HMI tags "DB_SDC_ERROR_STAT_EMS052"
   "DB_SDC_ERRORS_STAT_ER_AKT[52].ER_TRIGER" : Word = PLC DB_SDC_ERRORS_STAT.ER_AKT[52].ER_TRIGER AT %DB3724.DBW31386, 1 s
   "DB_SDC_ERRORS_STAT_ER_AKT[52].ER_STAT[1].DRIVE_POS" : DInt = PLC DB_SDC_ERRORS_STAT.ER_AKT[52].ER_STAT[1].DRIVE_POS AT %DB3724.DBD31392, 1 s
   "DB_SDC_ERRORS_STAT_ER_AKT[52].ER_STAT[1].ERROR" : Int = PLC DB_SDC_ERRORS_STAT.ER_AKT[52].ER_STAT[1].ERROR AT %DB3724.DBW31398, 1 s
   "DB_SDC_ERRORS_STAT_ER_AKT[52].ER_STAT[2].DRIVE_POS" : DInt = PLC DB_SDC_ERRORS_STAT.ER_AKT[52].ER_STAT[2].DRIVE_POS AT %DB3724.DBD31408, 1 s
   "DB_SDC_ERRORS_STAT_ER_AKT[52].ER_STAT[2].ERROR" : Int = PLC DB_SDC_ERRORS_STAT.ER_AKT[52].ER_STAT[2].ERROR AT %DB3724.DBW31414, 1 s
   "DB_SDC_ERRORS_STAT_ER_AKT[52].ER_STAT[3].DRIVE_POS" : DInt = PLC DB_SDC_ERRORS_STAT.ER_AKT[52].ER_STAT[3].DRIVE_POS AT %DB3724.DBD31424, 1 s
   "DB_SDC_ERRORS_STAT_ER_AKT[52].ER_STAT[3].ERROR" : Int = PLC DB_SDC_ERRORS_STAT.ER_AKT[52].ER_STAT[3].ERROR AT %DB3724.DBW31430, 1 s
   "DB_SDC_ERRORS_STAT_ER_AKT[52].ER_STAT[4].DRIVE_POS" : DInt = PLC DB_SDC_ERRORS_STAT.ER_AKT[52].ER_STAT[4].DRIVE_POS AT %DB3724.DBD31440, 1 s
   "DB_SDC_ERRORS_STAT_ER_AKT[52].ER_STAT[4].ERROR" : Int = PLC DB_SDC_ERRORS_STAT.ER_AKT[52].ER_STAT[4].ERROR AT %DB3724.DBW31446, 1 s

HMI tags "DB_SDC_ERROR_STAT_EMS053"
   "DB_SDC_ERRORS_STAT_ER_AKT[53].ER_TRIGER" : Word = PLC DB_SDC_ERRORS_STAT.ER_AKT[53].ER_TRIGER AT %DB3724.DBW31452, 1 s
   "DB_SDC_ERRORS_STAT_ER_AKT[53].ER_STAT[1].DRIVE_POS" : DInt = PLC DB_SDC_ERRORS_STAT.ER_AKT[53].ER_STAT[1].DRIVE_POS AT %DB3724.DBD31458, 1 s
   "DB_SDC_ERRORS_STAT_ER_AKT[53].ER_STAT[1].ERROR" : Int = PLC DB_SDC_ERRORS_STAT.ER_AKT[53].ER_STAT[1].ERROR AT %DB3724.DBW31464, 1 s
   "DB_SDC_ERRORS_STAT_ER_AKT[53].ER_STAT[2].DRIVE_POS" : DInt = PLC DB_SDC_ERRORS_STAT.ER_AKT[53].ER_STAT[2].DRIVE_POS AT %DB3724.DBD31474, 1 s
   "DB_SDC_ERRORS_STAT_ER_AKT[53].ER_STAT[2].ERROR" : Int = PLC DB_SDC_ERRORS_STAT.ER_AKT[53].ER_STAT[2].ERROR AT %DB3724.DBW31480, 1 s
   "DB_SDC_ERRORS_STAT_ER_AKT[53].ER_STAT[3].DRIVE_POS" : DInt = PLC DB_SDC_ERRORS_STAT.ER_AKT[53].ER_STAT[3].DRIVE_POS AT %DB3724.DBD31490, 1 s
   "DB_SDC_ERRORS_STAT_ER_AKT[53].ER_STAT[3].ERROR" : Int = PLC DB_SDC_ERRORS_STAT.ER_AKT[53].ER_STAT[3].ERROR AT %DB3724.DBW31496, 1 s
   "DB_SDC_ERRORS_STAT_ER_AKT[53].ER_STAT[4].DRIVE_POS" : DInt = PLC DB_SDC_ERRORS_STAT.ER_AKT[53].ER_STAT[4].DRIVE_POS AT %DB3724.DBD31506, 1 s
   "DB_SDC_ERRORS_STAT_ER_AKT[53].ER_STAT[4].ERROR" : Int = PLC DB_SDC_ERRORS_STAT.ER_AKT[53].ER_STAT[4].ERROR AT %DB3724.DBW31512, 1 s

HMI tags "DB_SDC_ERROR_STAT_EMS054"
   "DB_SDC_ERRORS_STAT_ER_AKT[54].ER_TRIGER" : Word = PLC DB_SDC_ERRORS_STAT.ER_AKT[54].ER_TRIGER AT %DB3724.DBW31518, 1 s
   "DB_SDC_ERRORS_STAT_ER_AKT[54].ER_STAT[1].DRIVE_POS" : DInt = PLC DB_SDC_ERRORS_STAT.ER_AKT[54].ER_STAT[1].DRIVE_POS AT %DB3724.DBD31524, 1 s
   "DB_SDC_ERRORS_STAT_ER_AKT[54].ER_STAT[1].ERROR" : Int = PLC DB_SDC_ERRORS_STAT.ER_AKT[54].ER_STAT[1].ERROR AT %DB3724.DBW31530, 1 s
   "DB_SDC_ERRORS_STAT_ER_AKT[54].ER_STAT[2].DRIVE_POS" : DInt = PLC DB_SDC_ERRORS_STAT.ER_AKT[54].ER_STAT[2].DRIVE_POS AT %DB3724.DBD31540, 1 s
   "DB_SDC_ERRORS_STAT_ER_AKT[54].ER_STAT[2].ERROR" : Int = PLC DB_SDC_ERRORS_STAT.ER_AKT[54].ER_STAT[2].ERROR AT %DB3724.DBW31546, 1 s
   "DB_SDC_ERRORS_STAT_ER_AKT[54].ER_STAT[3].DRIVE_POS" : DInt = PLC DB_SDC_ERRORS_STAT.ER_AKT[54].ER_STAT[3].DRIVE_POS AT %DB3724.DBD31556, 1 s
   "DB_SDC_ERRORS_STAT_ER_AKT[54].ER_STAT[3].ERROR" : Int = PLC DB_SDC_ERRORS_STAT.ER_AKT[54].ER_STAT[3].ERROR AT %DB3724.DBW31562, 1 s
   "DB_SDC_ERRORS_STAT_ER_AKT[54].ER_STAT[4].DRIVE_POS" : DInt = PLC DB_SDC_ERRORS_STAT.ER_AKT[54].ER_STAT[4].DRIVE_POS AT %DB3724.DBD31572, 1 s
   "DB_SDC_ERRORS_STAT_ER_AKT[54].ER_STAT[4].ERROR" : Int = PLC DB_SDC_ERRORS_STAT.ER_AKT[54].ER_STAT[4].ERROR AT %DB3724.DBW31578, 1 s

HMI tags "DB_SDC_ERROR_STAT_EMS055"
   "DB_SDC_ERRORS_STAT_ER_AKT[55].ER_TRIGER" : Word = PLC DB_SDC_ERRORS_STAT.ER_AKT[55].ER_TRIGER AT %DB3724.DBW31584, 1 s
   "DB_SDC_ERRORS_STAT_ER_AKT[55].ER_STAT[1].DRIVE_POS" : DInt = PLC DB_SDC_ERRORS_STAT.ER_AKT[55].ER_STAT[1].DRIVE_POS AT %DB3724.DBD31590, 1 s
   "DB_SDC_ERRORS_STAT_ER_AKT[55].ER_STAT[1].ERROR" : Int = PLC DB_SDC_ERRORS_STAT.ER_AKT[55].ER_STAT[1].ERROR AT %DB3724.DBW31596, 1 s
   "DB_SDC_ERRORS_STAT_ER_AKT[55].ER_STAT[2].DRIVE_POS" : DInt = PLC DB_SDC_ERRORS_STAT.ER_AKT[55].ER_STAT[2].DRIVE_POS AT %DB3724.DBD31606, 1 s
   "DB_SDC_ERRORS_STAT_ER_AKT[55].ER_STAT[2].ERROR" : Int = PLC DB_SDC_ERRORS_STAT.ER_AKT[55].ER_STAT[2].ERROR AT %DB3724.DBW31612, 1 s
   "DB_SDC_ERRORS_STAT_ER_AKT[55].ER_STAT[3].DRIVE_POS" : DInt = PLC DB_SDC_ERRORS_STAT.ER_AKT[55].ER_STAT[3].DRIVE_POS AT %DB3724.DBD31622, 1 s
   "DB_SDC_ERRORS_STAT_ER_AKT[55].ER_STAT[3].ERROR" : Int = PLC DB_SDC_ERRORS_STAT.ER_AKT[55].ER_STAT[3].ERROR AT %DB3724.DBW31628, 1 s
   "DB_SDC_ERRORS_STAT_ER_AKT[55].ER_STAT[4].DRIVE_POS" : DInt = PLC DB_SDC_ERRORS_STAT.ER_AKT[55].ER_STAT[4].DRIVE_POS AT %DB3724.DBD31638, 1 s
   "DB_SDC_ERRORS_STAT_ER_AKT[55].ER_STAT[4].ERROR" : Int = PLC DB_SDC_ERRORS_STAT.ER_AKT[55].ER_STAT[4].ERROR AT %DB3724.DBW31644, 1 s

HMI tags "DB_SDC_ERROR_STAT_EMS056"
   "DB_SDC_ERRORS_STAT_ER_AKT[56].ER_TRIGER" : Word = PLC DB_SDC_ERRORS_STAT.ER_AKT[56].ER_TRIGER AT %DB3724.DBW31650, 1 s
   "DB_SDC_ERRORS_STAT_ER_AKT[56].ER_STAT[1].DRIVE_POS" : DInt = PLC DB_SDC_ERRORS_STAT.ER_AKT[56].ER_STAT[1].DRIVE_POS AT %DB3724.DBD31656, 1 s
   "DB_SDC_ERRORS_STAT_ER_AKT[56].ER_STAT[1].ERROR" : Int = PLC DB_SDC_ERRORS_STAT.ER_AKT[56].ER_STAT[1].ERROR AT %DB3724.DBW31662, 1 s
   "DB_SDC_ERRORS_STAT_ER_AKT[56].ER_STAT[2].DRIVE_POS" : DInt = PLC DB_SDC_ERRORS_STAT.ER_AKT[56].ER_STAT[2].DRIVE_POS AT %DB3724.DBD31672, 1 s
   "DB_SDC_ERRORS_STAT_ER_AKT[56].ER_STAT[2].ERROR" : Int = PLC DB_SDC_ERRORS_STAT.ER_AKT[56].ER_STAT[2].ERROR AT %DB3724.DBW31678, 1 s
   "DB_SDC_ERRORS_STAT_ER_AKT[56].ER_STAT[3].DRIVE_POS" : DInt = PLC DB_SDC_ERRORS_STAT.ER_AKT[56].ER_STAT[3].DRIVE_POS AT %DB3724.DBD31688, 1 s
   "DB_SDC_ERRORS_STAT_ER_AKT[56].ER_STAT[3].ERROR" : Int = PLC DB_SDC_ERRORS_STAT.ER_AKT[56].ER_STAT[3].ERROR AT %DB3724.DBW31694, 1 s
   "DB_SDC_ERRORS_STAT_ER_AKT[56].ER_STAT[4].DRIVE_POS" : DInt = PLC DB_SDC_ERRORS_STAT.ER_AKT[56].ER_STAT[4].DRIVE_POS AT %DB3724.DBD31704, 1 s
   "DB_SDC_ERRORS_STAT_ER_AKT[56].ER_STAT[4].ERROR" : Int = PLC DB_SDC_ERRORS_STAT.ER_AKT[56].ER_STAT[4].ERROR AT %DB3724.DBW31710, 1 s

HMI tags "DB_SDC_ERROR_STAT_EMS057"
   "DB_SDC_ERRORS_STAT_ER_AKT[57].ER_TRIGER" : Word = PLC DB_SDC_ERRORS_STAT.ER_AKT[57].ER_TRIGER AT %DB3724.DBW31716, 1 s
   "DB_SDC_ERRORS_STAT_ER_AKT[57].ER_STAT[1].DRIVE_POS" : DInt = PLC DB_SDC_ERRORS_STAT.ER_AKT[57].ER_STAT[1].DRIVE_POS AT %DB3724.DBD31722, 1 s
   "DB_SDC_ERRORS_STAT_ER_AKT[57].ER_STAT[1].ERROR" : Int = PLC DB_SDC_ERRORS_STAT.ER_AKT[57].ER_STAT[1].ERROR AT %DB3724.DBW31728, 1 s
   "DB_SDC_ERRORS_STAT_ER_AKT[57].ER_STAT[2].DRIVE_POS" : DInt = PLC DB_SDC_ERRORS_STAT.ER_AKT[57].ER_STAT[2].DRIVE_POS AT %DB3724.DBD31738, 1 s
   "DB_SDC_ERRORS_STAT_ER_AKT[57].ER_STAT[2].ERROR" : Int = PLC DB_SDC_ERRORS_STAT.ER_AKT[57].ER_STAT[2].ERROR AT %DB3724.DBW31744, 1 s
   "DB_SDC_ERRORS_STAT_ER_AKT[57].ER_STAT[3].DRIVE_POS" : DInt = PLC DB_SDC_ERRORS_STAT.ER_AKT[57].ER_STAT[3].DRIVE_POS AT %DB3724.DBD31754, 1 s
   "DB_SDC_ERRORS_STAT_ER_AKT[57].ER_STAT[3].ERROR" : Int = PLC DB_SDC_ERRORS_STAT.ER_AKT[57].ER_STAT[3].ERROR AT %DB3724.DBW31760, 1 s
   "DB_SDC_ERRORS_STAT_ER_AKT[57].ER_STAT[4].DRIVE_POS" : DInt = PLC DB_SDC_ERRORS_STAT.ER_AKT[57].ER_STAT[4].DRIVE_POS AT %DB3724.DBD31770, 1 s
   "DB_SDC_ERRORS_STAT_ER_AKT[57].ER_STAT[4].ERROR" : Int = PLC DB_SDC_ERRORS_STAT.ER_AKT[57].ER_STAT[4].ERROR AT %DB3724.DBW31776, 1 s

HMI tags "DB_SDC_ERROR_STAT_EMS058"
   "DB_SDC_ERRORS_STAT_ER_AKT[58].ER_TRIGER" : Word = PLC DB_SDC_ERRORS_STAT.ER_AKT[58].ER_TRIGER AT %DB3724.DBW31782, 1 s
   "DB_SDC_ERRORS_STAT_ER_AKT[58].ER_STAT[1].DRIVE_POS" : DInt = PLC DB_SDC_ERRORS_STAT.ER_AKT[58].ER_STAT[1].DRIVE_POS AT %DB3724.DBD31788, 1 s
   "DB_SDC_ERRORS_STAT_ER_AKT[58].ER_STAT[1].ERROR" : Int = PLC DB_SDC_ERRORS_STAT.ER_AKT[58].ER_STAT[1].ERROR AT %DB3724.DBW31794, 1 s
   "DB_SDC_ERRORS_STAT_ER_AKT[58].ER_STAT[2].DRIVE_POS" : DInt = PLC DB_SDC_ERRORS_STAT.ER_AKT[58].ER_STAT[2].DRIVE_POS AT %DB3724.DBD31804, 1 s
   "DB_SDC_ERRORS_STAT_ER_AKT[58].ER_STAT[2].ERROR" : Int = PLC DB_SDC_ERRORS_STAT.ER_AKT[58].ER_STAT[2].ERROR AT %DB3724.DBW31810, 1 s
   "DB_SDC_ERRORS_STAT_ER_AKT[58].ER_STAT[3].DRIVE_POS" : DInt = PLC DB_SDC_ERRORS_STAT.ER_AKT[58].ER_STAT[3].DRIVE_POS AT %DB3724.DBD31820, 1 s
   "DB_SDC_ERRORS_STAT_ER_AKT[58].ER_STAT[3].ERROR" : Int = PLC DB_SDC_ERRORS_STAT.ER_AKT[58].ER_STAT[3].ERROR AT %DB3724.DBW31826, 1 s
   "DB_SDC_ERRORS_STAT_ER_AKT[58].ER_STAT[4].DRIVE_POS" : DInt = PLC DB_SDC_ERRORS_STAT.ER_AKT[58].ER_STAT[4].DRIVE_POS AT %DB3724.DBD31836, 1 s
   "DB_SDC_ERRORS_STAT_ER_AKT[58].ER_STAT[4].ERROR" : Int = PLC DB_SDC_ERRORS_STAT.ER_AKT[58].ER_STAT[4].ERROR AT %DB3724.DBW31842, 1 s

HMI tags "DB_SDC_ERROR_STAT_EMS059"
   "DB_SDC_ERRORS_STAT_ER_AKT[59].ER_TRIGER" : Word = PLC DB_SDC_ERRORS_STAT.ER_AKT[59].ER_TRIGER AT %DB3724.DBW31848, 1 s
   "DB_SDC_ERRORS_STAT_ER_AKT[59].ER_STAT[1].DRIVE_POS" : DInt = PLC DB_SDC_ERRORS_STAT.ER_AKT[59].ER_STAT[1].DRIVE_POS AT %DB3724.DBD31854, 1 s
   "DB_SDC_ERRORS_STAT_ER_AKT[59].ER_STAT[1].ERROR" : Int = PLC DB_SDC_ERRORS_STAT.ER_AKT[59].ER_STAT[1].ERROR AT %DB3724.DBW31860, 1 s
   "DB_SDC_ERRORS_STAT_ER_AKT[59].ER_STAT[2].DRIVE_POS" : DInt = PLC DB_SDC_ERRORS_STAT.ER_AKT[59].ER_STAT[2].DRIVE_POS AT %DB3724.DBD31870, 1 s
   "DB_SDC_ERRORS_STAT_ER_AKT[59].ER_STAT[2].ERROR" : Int = PLC DB_SDC_ERRORS_STAT.ER_AKT[59].ER_STAT[2].ERROR AT %DB3724.DBW31876, 1 s
   "DB_SDC_ERRORS_STAT_ER_AKT[59].ER_STAT[3].DRIVE_POS" : DInt = PLC DB_SDC_ERRORS_STAT.ER_AKT[59].ER_STAT[3].DRIVE_POS AT %DB3724.DBD31886, 1 s
   "DB_SDC_ERRORS_STAT_ER_AKT[59].ER_STAT[3].ERROR" : Int = PLC DB_SDC_ERRORS_STAT.ER_AKT[59].ER_STAT[3].ERROR AT %DB3724.DBW31892, 1 s
   "DB_SDC_ERRORS_STAT_ER_AKT[59].ER_STAT[4].DRIVE_POS" : DInt = PLC DB_SDC_ERRORS_STAT.ER_AKT[59].ER_STAT[4].DRIVE_POS AT %DB3724.DBD31902, 1 s
   "DB_SDC_ERRORS_STAT_ER_AKT[59].ER_STAT[4].ERROR" : Int = PLC DB_SDC_ERRORS_STAT.ER_AKT[59].ER_STAT[4].ERROR AT %DB3724.DBW31908, 1 s

HMI tags "DB_SDC_ERROR_STAT_EMS060"
   "DB_SDC_ERRORS_STAT_ER_AKT[60].ER_TRIGER" : Word = PLC DB_SDC_ERRORS_STAT.ER_AKT[60].ER_TRIGER AT %DB3724.DBW31914, 1 s
   "DB_SDC_ERRORS_STAT_ER_AKT[60].ER_STAT[1].DRIVE_POS" : DInt = PLC DB_SDC_ERRORS_STAT.ER_AKT[60].ER_STAT[1].DRIVE_POS AT %DB3724.DBD31920, 1 s
   "DB_SDC_ERRORS_STAT_ER_AKT[60].ER_STAT[1].ERROR" : Int = PLC DB_SDC_ERRORS_STAT.ER_AKT[60].ER_STAT[1].ERROR AT %DB3724.DBW31926, 1 s
   "DB_SDC_ERRORS_STAT_ER_AKT[60].ER_STAT[2].DRIVE_POS" : DInt = PLC DB_SDC_ERRORS_STAT.ER_AKT[60].ER_STAT[2].DRIVE_POS AT %DB3724.DBD31936, 1 s
   "DB_SDC_ERRORS_STAT_ER_AKT[60].ER_STAT[2].ERROR" : Int = PLC DB_SDC_ERRORS_STAT.ER_AKT[60].ER_STAT[2].ERROR AT %DB3724.DBW31942, 1 s
   "DB_SDC_ERRORS_STAT_ER_AKT[60].ER_STAT[3].DRIVE_POS" : DInt = PLC DB_SDC_ERRORS_STAT.ER_AKT[60].ER_STAT[3].DRIVE_POS AT %DB3724.DBD31952, 1 s
   "DB_SDC_ERRORS_STAT_ER_AKT[60].ER_STAT[3].ERROR" : Int = PLC DB_SDC_ERRORS_STAT.ER_AKT[60].ER_STAT[3].ERROR AT %DB3724.DBW31958, 1 s
   "DB_SDC_ERRORS_STAT_ER_AKT[60].ER_STAT[4].DRIVE_POS" : DInt = PLC DB_SDC_ERRORS_STAT.ER_AKT[60].ER_STAT[4].DRIVE_POS AT %DB3724.DBD31968, 1 s
   "DB_SDC_ERRORS_STAT_ER_AKT[60].ER_STAT[4].ERROR" : Int = PLC DB_SDC_ERRORS_STAT.ER_AKT[60].ER_STAT[4].ERROR AT %DB3724.DBW31974, 1 s

HMI tags "DB_SDC_ERROR_STAT_EMS061"
   "DB_SDC_ERRORS_STAT_ER_AKT[61].ER_TRIGER" : Word = PLC DB_SDC_ERRORS_STAT.ER_AKT[61].ER_TRIGER AT %DB3724.DBW31980, 1 s
   "DB_SDC_ERRORS_STAT_ER_AKT[61].ER_STAT[1].DRIVE_POS" : DInt = PLC DB_SDC_ERRORS_STAT.ER_AKT[61].ER_STAT[1].DRIVE_POS AT %DB3724.DBD31986, 1 s
   "DB_SDC_ERRORS_STAT_ER_AKT[61].ER_STAT[1].ERROR" : Int = PLC DB_SDC_ERRORS_STAT.ER_AKT[61].ER_STAT[1].ERROR AT %DB3724.DBW31992, 1 s
   "DB_SDC_ERRORS_STAT_ER_AKT[61].ER_STAT[2].DRIVE_POS" : DInt = PLC DB_SDC_ERRORS_STAT.ER_AKT[61].ER_STAT[2].DRIVE_POS AT %DB3724.DBD32002, 1 s
   "DB_SDC_ERRORS_STAT_ER_AKT[61].ER_STAT[2].ERROR" : Int = PLC DB_SDC_ERRORS_STAT.ER_AKT[61].ER_STAT[2].ERROR AT %DB3724.DBW32008, 1 s
   "DB_SDC_ERRORS_STAT_ER_AKT[61].ER_STAT[3].DRIVE_POS" : DInt = PLC DB_SDC_ERRORS_STAT.ER_AKT[61].ER_STAT[3].DRIVE_POS AT %DB3724.DBD32018, 1 s
   "DB_SDC_ERRORS_STAT_ER_AKT[61].ER_STAT[3].ERROR" : Int = PLC DB_SDC_ERRORS_STAT.ER_AKT[61].ER_STAT[3].ERROR AT %DB3724.DBW32024, 1 s
   "DB_SDC_ERRORS_STAT_ER_AKT[61].ER_STAT[4].DRIVE_POS" : DInt = PLC DB_SDC_ERRORS_STAT.ER_AKT[61].ER_STAT[4].DRIVE_POS AT %DB3724.DBD32034, 1 s
   "DB_SDC_ERRORS_STAT_ER_AKT[61].ER_STAT[4].ERROR" : Int = PLC DB_SDC_ERRORS_STAT.ER_AKT[61].ER_STAT[4].ERROR AT %DB3724.DBW32040, 1 s

HMI tags "DB_SDC_ERROR_STAT_EMS062"
   "DB_SDC_ERRORS_STAT_ER_AKT[62].ER_TRIGER" : Word = PLC DB_SDC_ERRORS_STAT.ER_AKT[62].ER_TRIGER AT %DB3724.DBW32046, 1 s
   "DB_SDC_ERRORS_STAT_ER_AKT[62].ER_STAT[1].DRIVE_POS" : DInt = PLC DB_SDC_ERRORS_STAT.ER_AKT[62].ER_STAT[1].DRIVE_POS AT %DB3724.DBD32052, 1 s
   "DB_SDC_ERRORS_STAT_ER_AKT[62].ER_STAT[1].ERROR" : Int = PLC DB_SDC_ERRORS_STAT.ER_AKT[62].ER_STAT[1].ERROR AT %DB3724.DBW32058, 1 s
   "DB_SDC_ERRORS_STAT_ER_AKT[62].ER_STAT[2].DRIVE_POS" : DInt = PLC DB_SDC_ERRORS_STAT.ER_AKT[62].ER_STAT[2].DRIVE_POS AT %DB3724.DBD32068, 1 s
   "DB_SDC_ERRORS_STAT_ER_AKT[62].ER_STAT[2].ERROR" : Int = PLC DB_SDC_ERRORS_STAT.ER_AKT[62].ER_STAT[2].ERROR AT %DB3724.DBW32074, 1 s
   "DB_SDC_ERRORS_STAT_ER_AKT[62].ER_STAT[3].DRIVE_POS" : DInt = PLC DB_SDC_ERRORS_STAT.ER_AKT[62].ER_STAT[3].DRIVE_POS AT %DB3724.DBD32084, 1 s
   "DB_SDC_ERRORS_STAT_ER_AKT[62].ER_STAT[3].ERROR" : Int = PLC DB_SDC_ERRORS_STAT.ER_AKT[62].ER_STAT[3].ERROR AT %DB3724.DBW32090, 1 s
   "DB_SDC_ERRORS_STAT_ER_AKT[62].ER_STAT[4].DRIVE_POS" : DInt = PLC DB_SDC_ERRORS_STAT.ER_AKT[62].ER_STAT[4].DRIVE_POS AT %DB3724.DBD32100, 1 s
   "DB_SDC_ERRORS_STAT_ER_AKT[62].ER_STAT[4].ERROR" : Int = PLC DB_SDC_ERRORS_STAT.ER_AKT[62].ER_STAT[4].ERROR AT %DB3724.DBW32106, 1 s

HMI tags "DB_SDC_ERROR_STAT_EMS063"
   "DB_SDC_ERRORS_STAT_ER_AKT[63].ER_TRIGER" : Word = PLC DB_SDC_ERRORS_STAT.ER_AKT[63].ER_TRIGER AT %DB3724.DBW32112, 1 s
   "DB_SDC_ERRORS_STAT_ER_AKT[63].ER_STAT[1].DRIVE_POS" : DInt = PLC DB_SDC_ERRORS_STAT.ER_AKT[63].ER_STAT[1].DRIVE_POS AT %DB3724.DBD32118, 1 s
   "DB_SDC_ERRORS_STAT_ER_AKT[63].ER_STAT[1].ERROR" : Int = PLC DB_SDC_ERRORS_STAT.ER_AKT[63].ER_STAT[1].ERROR AT %DB3724.DBW32124, 1 s
   "DB_SDC_ERRORS_STAT_ER_AKT[63].ER_STAT[2].DRIVE_POS" : DInt = PLC DB_SDC_ERRORS_STAT.ER_AKT[63].ER_STAT[2].DRIVE_POS AT %DB3724.DBD32134, 1 s
   "DB_SDC_ERRORS_STAT_ER_AKT[63].ER_STAT[2].ERROR" : Int = PLC DB_SDC_ERRORS_STAT.ER_AKT[63].ER_STAT[2].ERROR AT %DB3724.DBW32140, 1 s
   "DB_SDC_ERRORS_STAT_ER_AKT[63].ER_STAT[3].DRIVE_POS" : DInt = PLC DB_SDC_ERRORS_STAT.ER_AKT[63].ER_STAT[3].DRIVE_POS AT %DB3724.DBD32150, 1 s
   "DB_SDC_ERRORS_STAT_ER_AKT[63].ER_STAT[3].ERROR" : Int = PLC DB_SDC_ERRORS_STAT.ER_AKT[63].ER_STAT[3].ERROR AT %DB3724.DBW32156, 1 s
   "DB_SDC_ERRORS_STAT_ER_AKT[63].ER_STAT[4].DRIVE_POS" : DInt = PLC DB_SDC_ERRORS_STAT.ER_AKT[63].ER_STAT[4].DRIVE_POS AT %DB3724.DBD32166, 1 s
   "DB_SDC_ERRORS_STAT_ER_AKT[63].ER_STAT[4].ERROR" : Int = PLC DB_SDC_ERRORS_STAT.ER_AKT[63].ER_STAT[4].ERROR AT %DB3724.DBW32172, 1 s

HMI tags "DB_SDC_ERROR_STAT_EMS064"
   "DB_SDC_ERRORS_STAT_ER_AKT[64].ER_TRIGER" : Word = PLC DB_SDC_ERRORS_STAT.ER_AKT[64].ER_TRIGER AT %DB3724.DBW32178, 1 s
   "DB_SDC_ERRORS_STAT_ER_AKT[64].ER_STAT[1].DRIVE_POS" : DInt = PLC DB_SDC_ERRORS_STAT.ER_AKT[64].ER_STAT[1].DRIVE_POS AT %DB3724.DBD32184, 1 s
   "DB_SDC_ERRORS_STAT_ER_AKT[64].ER_STAT[1].ERROR" : Int = PLC DB_SDC_ERRORS_STAT.ER_AKT[64].ER_STAT[1].ERROR AT %DB3724.DBW32190, 1 s
   "DB_SDC_ERRORS_STAT_ER_AKT[64].ER_STAT[2].DRIVE_POS" : DInt = PLC DB_SDC_ERRORS_STAT.ER_AKT[64].ER_STAT[2].DRIVE_POS AT %DB3724.DBD32200, 1 s
   "DB_SDC_ERRORS_STAT_ER_AKT[64].ER_STAT[2].ERROR" : Int = PLC DB_SDC_ERRORS_STAT.ER_AKT[64].ER_STAT[2].ERROR AT %DB3724.DBW32206, 1 s
   "DB_SDC_ERRORS_STAT_ER_AKT[64].ER_STAT[3].DRIVE_POS" : DInt = PLC DB_SDC_ERRORS_STAT.ER_AKT[64].ER_STAT[3].DRIVE_POS AT %DB3724.DBD32216, 1 s
   "DB_SDC_ERRORS_STAT_ER_AKT[64].ER_STAT[3].ERROR" : Int = PLC DB_SDC_ERRORS_STAT.ER_AKT[64].ER_STAT[3].ERROR AT %DB3724.DBW32222, 1 s
   "DB_SDC_ERRORS_STAT_ER_AKT[64].ER_STAT[4].DRIVE_POS" : DInt = PLC DB_SDC_ERRORS_STAT.ER_AKT[64].ER_STAT[4].DRIVE_POS AT %DB3724.DBD32232, 1 s
   "DB_SDC_ERRORS_STAT_ER_AKT[64].ER_STAT[4].ERROR" : Int = PLC DB_SDC_ERRORS_STAT.ER_AKT[64].ER_STAT[4].ERROR AT %DB3724.DBW32238, 1 s

HMI tags "DB_SDC_ERROR_STAT_EMS065"
   "DB_SDC_ERRORS_STAT_ER_AKT[65].ER_TRIGER" : Word = PLC DB_SDC_ERRORS_STAT.ER_AKT[65].ER_TRIGER AT %DB3724.DBW32244, 1 s
   "DB_SDC_ERRORS_STAT_ER_AKT[65].ER_STAT[1].DRIVE_POS" : DInt = PLC DB_SDC_ERRORS_STAT.ER_AKT[65].ER_STAT[1].DRIVE_POS AT %DB3724.DBD32250, 1 s
   "DB_SDC_ERRORS_STAT_ER_AKT[65].ER_STAT[1].ERROR" : Int = PLC DB_SDC_ERRORS_STAT.ER_AKT[65].ER_STAT[1].ERROR AT %DB3724.DBW32256, 1 s
   "DB_SDC_ERRORS_STAT_ER_AKT[65].ER_STAT[2].DRIVE_POS" : DInt = PLC DB_SDC_ERRORS_STAT.ER_AKT[65].ER_STAT[2].DRIVE_POS AT %DB3724.DBD32266, 1 s
   "DB_SDC_ERRORS_STAT_ER_AKT[65].ER_STAT[2].ERROR" : Int = PLC DB_SDC_ERRORS_STAT.ER_AKT[65].ER_STAT[2].ERROR AT %DB3724.DBW32272, 1 s
   "DB_SDC_ERRORS_STAT_ER_AKT[65].ER_STAT[3].DRIVE_POS" : DInt = PLC DB_SDC_ERRORS_STAT.ER_AKT[65].ER_STAT[3].DRIVE_POS AT %DB3724.DBD32282, 1 s
   "DB_SDC_ERRORS_STAT_ER_AKT[65].ER_STAT[3].ERROR" : Int = PLC DB_SDC_ERRORS_STAT.ER_AKT[65].ER_STAT[3].ERROR AT %DB3724.DBW32288, 1 s
   "DB_SDC_ERRORS_STAT_ER_AKT[65].ER_STAT[4].DRIVE_POS" : DInt = PLC DB_SDC_ERRORS_STAT.ER_AKT[65].ER_STAT[4].DRIVE_POS AT %DB3724.DBD32298, 1 s
   "DB_SDC_ERRORS_STAT_ER_AKT[65].ER_STAT[4].ERROR" : Int = PLC DB_SDC_ERRORS_STAT.ER_AKT[65].ER_STAT[4].ERROR AT %DB3724.DBW32304, 1 s

HMI tags "DB_SDC_ERROR_STAT_EMS066"
   "DB_SDC_ERRORS_STAT_ER_AKT[66].ER_TRIGER" : Word = PLC DB_SDC_ERRORS_STAT.ER_AKT[66].ER_TRIGER AT %DB3724.DBW32310, 1 s
   "DB_SDC_ERRORS_STAT_ER_AKT[66].ER_STAT[1].DRIVE_POS" : DInt = PLC DB_SDC_ERRORS_STAT.ER_AKT[66].ER_STAT[1].DRIVE_POS AT %DB3724.DBD32316, 1 s
   "DB_SDC_ERRORS_STAT_ER_AKT[66].ER_STAT[1].ERROR" : Int = PLC DB_SDC_ERRORS_STAT.ER_AKT[66].ER_STAT[1].ERROR AT %DB3724.DBW32322, 1 s
   "DB_SDC_ERRORS_STAT_ER_AKT[66].ER_STAT[2].DRIVE_POS" : DInt = PLC DB_SDC_ERRORS_STAT.ER_AKT[66].ER_STAT[2].DRIVE_POS AT %DB3724.DBD32332, 1 s
   "DB_SDC_ERRORS_STAT_ER_AKT[66].ER_STAT[2].ERROR" : Int = PLC DB_SDC_ERRORS_STAT.ER_AKT[66].ER_STAT[2].ERROR AT %DB3724.DBW32338, 1 s
   "DB_SDC_ERRORS_STAT_ER_AKT[66].ER_STAT[3].DRIVE_POS" : DInt = PLC DB_SDC_ERRORS_STAT.ER_AKT[66].ER_STAT[3].DRIVE_POS AT %DB3724.DBD32348, 1 s
   "DB_SDC_ERRORS_STAT_ER_AKT[66].ER_STAT[3].ERROR" : Int = PLC DB_SDC_ERRORS_STAT.ER_AKT[66].ER_STAT[3].ERROR AT %DB3724.DBW32354, 1 s
   "DB_SDC_ERRORS_STAT_ER_AKT[66].ER_STAT[4].DRIVE_POS" : DInt = PLC DB_SDC_ERRORS_STAT.ER_AKT[66].ER_STAT[4].DRIVE_POS AT %DB3724.DBD32364, 1 s
   "DB_SDC_ERRORS_STAT_ER_AKT[66].ER_STAT[4].ERROR" : Int = PLC DB_SDC_ERRORS_STAT.ER_AKT[66].ER_STAT[4].ERROR AT %DB3724.DBW32370, 1 s

HMI tags "DB_SDC_ERROR_STAT_EMS067"
   "DB_SDC_ERRORS_STAT_ER_AKT[67].ER_TRIGER" : Word = PLC DB_SDC_ERRORS_STAT.ER_AKT[67].ER_TRIGER AT %DB3724.DBW32376, 1 s
   "DB_SDC_ERRORS_STAT_ER_AKT[67].ER_STAT[1].DRIVE_POS" : DInt = PLC DB_SDC_ERRORS_STAT.ER_AKT[67].ER_STAT[1].DRIVE_POS AT %DB3724.DBD32382, 1 s
   "DB_SDC_ERRORS_STAT_ER_AKT[67].ER_STAT[1].ERROR" : Int = PLC DB_SDC_ERRORS_STAT.ER_AKT[67].ER_STAT[1].ERROR AT %DB3724.DBW32388, 1 s
   "DB_SDC_ERRORS_STAT_ER_AKT[67].ER_STAT[2].DRIVE_POS" : DInt = PLC DB_SDC_ERRORS_STAT.ER_AKT[67].ER_STAT[2].DRIVE_POS AT %DB3724.DBD32398, 1 s
   "DB_SDC_ERRORS_STAT_ER_AKT[67].ER_STAT[2].ERROR" : Int = PLC DB_SDC_ERRORS_STAT.ER_AKT[67].ER_STAT[2].ERROR AT %DB3724.DBW32404, 1 s
   "DB_SDC_ERRORS_STAT_ER_AKT[67].ER_STAT[3].DRIVE_POS" : DInt = PLC DB_SDC_ERRORS_STAT.ER_AKT[67].ER_STAT[3].DRIVE_POS AT %DB3724.DBD32414, 1 s
   "DB_SDC_ERRORS_STAT_ER_AKT[67].ER_STAT[3].ERROR" : Int = PLC DB_SDC_ERRORS_STAT.ER_AKT[67].ER_STAT[3].ERROR AT %DB3724.DBW32420, 1 s
   "DB_SDC_ERRORS_STAT_ER_AKT[67].ER_STAT[4].DRIVE_POS" : DInt = PLC DB_SDC_ERRORS_STAT.ER_AKT[67].ER_STAT[4].DRIVE_POS AT %DB3724.DBD32430, 1 s
   "DB_SDC_ERRORS_STAT_ER_AKT[67].ER_STAT[4].ERROR" : Int = PLC DB_SDC_ERRORS_STAT.ER_AKT[67].ER_STAT[4].ERROR AT %DB3724.DBW32436, 1 s

HMI tags "DB_SDC_ERROR_STAT_EMS068"
   "DB_SDC_ERRORS_STAT_ER_AKT[68].ER_TRIGER" : Word = PLC DB_SDC_ERRORS_STAT.ER_AKT[68].ER_TRIGER AT %DB3724.DBW32442, 1 s
   "DB_SDC_ERRORS_STAT_ER_AKT[68].ER_STAT[1].DRIVE_POS" : DInt = PLC DB_SDC_ERRORS_STAT.ER_AKT[68].ER_STAT[1].DRIVE_POS AT %DB3724.DBD32448, 1 s
   "DB_SDC_ERRORS_STAT_ER_AKT[68].ER_STAT[1].ERROR" : Int = PLC DB_SDC_ERRORS_STAT.ER_AKT[68].ER_STAT[1].ERROR AT %DB3724.DBW32454, 1 s
   "DB_SDC_ERRORS_STAT_ER_AKT[68].ER_STAT[2].DRIVE_POS" : DInt = PLC DB_SDC_ERRORS_STAT.ER_AKT[68].ER_STAT[2].DRIVE_POS AT %DB3724.DBD32464, 1 s
   "DB_SDC_ERRORS_STAT_ER_AKT[68].ER_STAT[2].ERROR" : Int = PLC DB_SDC_ERRORS_STAT.ER_AKT[68].ER_STAT[2].ERROR AT %DB3724.DBW32470, 1 s
   "DB_SDC_ERRORS_STAT_ER_AKT[68].ER_STAT[3].DRIVE_POS" : DInt = PLC DB_SDC_ERRORS_STAT.ER_AKT[68].ER_STAT[3].DRIVE_POS AT %DB3724.DBD32480, 1 s
   "DB_SDC_ERRORS_STAT_ER_AKT[68].ER_STAT[3].ERROR" : Int = PLC DB_SDC_ERRORS_STAT.ER_AKT[68].ER_STAT[3].ERROR AT %DB3724.DBW32486, 1 s
   "DB_SDC_ERRORS_STAT_ER_AKT[68].ER_STAT[4].DRIVE_POS" : DInt = PLC DB_SDC_ERRORS_STAT.ER_AKT[68].ER_STAT[4].DRIVE_POS AT %DB3724.DBD32496, 1 s
   "DB_SDC_ERRORS_STAT_ER_AKT[68].ER_STAT[4].ERROR" : Int = PLC DB_SDC_ERRORS_STAT.ER_AKT[68].ER_STAT[4].ERROR AT %DB3724.DBW32502, 1 s

HMI tags "DB_SDC_ERROR_STAT_EMS069"
   "DB_SDC_ERRORS_STAT_ER_AKT[69].ER_TRIGER" : Word = PLC DB_SDC_ERRORS_STAT.ER_AKT[69].ER_TRIGER AT %DB3724.DBW32508, 1 s
   "DB_SDC_ERRORS_STAT_ER_AKT[69].ER_STAT[1].DRIVE_POS" : DInt = PLC DB_SDC_ERRORS_STAT.ER_AKT[69].ER_STAT[1].DRIVE_POS AT %DB3724.DBD32514, 1 s
   "DB_SDC_ERRORS_STAT_ER_AKT[69].ER_STAT[1].ERROR" : Int = PLC DB_SDC_ERRORS_STAT.ER_AKT[69].ER_STAT[1].ERROR AT %DB3724.DBW32520, 1 s
   "DB_SDC_ERRORS_STAT_ER_AKT[69].ER_STAT[2].DRIVE_POS" : DInt = PLC DB_SDC_ERRORS_STAT.ER_AKT[69].ER_STAT[2].DRIVE_POS AT %DB3724.DBD32530, 1 s
   "DB_SDC_ERRORS_STAT_ER_AKT[69].ER_STAT[2].ERROR" : Int = PLC DB_SDC_ERRORS_STAT.ER_AKT[69].ER_STAT[2].ERROR AT %DB3724.DBW32536, 1 s
   "DB_SDC_ERRORS_STAT_ER_AKT[69].ER_STAT[3].DRIVE_POS" : DInt = PLC DB_SDC_ERRORS_STAT.ER_AKT[69].ER_STAT[3].DRIVE_POS AT %DB3724.DBD32546, 1 s
   "DB_SDC_ERRORS_STAT_ER_AKT[69].ER_STAT[3].ERROR" : Int = PLC DB_SDC_ERRORS_STAT.ER_AKT[69].ER_STAT[3].ERROR AT %DB3724.DBW32552, 1 s
   "DB_SDC_ERRORS_STAT_ER_AKT[69].ER_STAT[4].DRIVE_POS" : DInt = PLC DB_SDC_ERRORS_STAT.ER_AKT[69].ER_STAT[4].DRIVE_POS AT %DB3724.DBD32562, 1 s
   "DB_SDC_ERRORS_STAT_ER_AKT[69].ER_STAT[4].ERROR" : Int = PLC DB_SDC_ERRORS_STAT.ER_AKT[69].ER_STAT[4].ERROR AT %DB3724.DBW32568, 1 s

HMI tags "DB_SDC_ERROR_STAT_EMS070"
   "DB_SDC_ERRORS_STAT_ER_AKT[70].ER_TRIGER" : Word = PLC DB_SDC_ERRORS_STAT.ER_AKT[70].ER_TRIGER AT %DB3724.DBW32574, 1 s
   "DB_SDC_ERRORS_STAT_ER_AKT[70].ER_STAT[1].DRIVE_POS" : DInt = PLC DB_SDC_ERRORS_STAT.ER_AKT[70].ER_STAT[1].DRIVE_POS AT %DB3724.DBD32580, 1 s
   "DB_SDC_ERRORS_STAT_ER_AKT[70].ER_STAT[1].ERROR" : Int = PLC DB_SDC_ERRORS_STAT.ER_AKT[70].ER_STAT[1].ERROR AT %DB3724.DBW32586, 1 s
   "DB_SDC_ERRORS_STAT_ER_AKT[70].ER_STAT[2].DRIVE_POS" : DInt = PLC DB_SDC_ERRORS_STAT.ER_AKT[70].ER_STAT[2].DRIVE_POS AT %DB3724.DBD32596, 1 s
   "DB_SDC_ERRORS_STAT_ER_AKT[70].ER_STAT[2].ERROR" : Int = PLC DB_SDC_ERRORS_STAT.ER_AKT[70].ER_STAT[2].ERROR AT %DB3724.DBW32602, 1 s
   "DB_SDC_ERRORS_STAT_ER_AKT[70].ER_STAT[3].DRIVE_POS" : DInt = PLC DB_SDC_ERRORS_STAT.ER_AKT[70].ER_STAT[3].DRIVE_POS AT %DB3724.DBD32612, 1 s
   "DB_SDC_ERRORS_STAT_ER_AKT[70].ER_STAT[3].ERROR" : Int = PLC DB_SDC_ERRORS_STAT.ER_AKT[70].ER_STAT[3].ERROR AT %DB3724.DBW32618, 1 s
   "DB_SDC_ERRORS_STAT_ER_AKT[70].ER_STAT[4].DRIVE_POS" : DInt = PLC DB_SDC_ERRORS_STAT.ER_AKT[70].ER_STAT[4].DRIVE_POS AT %DB3724.DBD32628, 1 s
   "DB_SDC_ERRORS_STAT_ER_AKT[70].ER_STAT[4].ERROR" : Int = PLC DB_SDC_ERRORS_STAT.ER_AKT[70].ER_STAT[4].ERROR AT %DB3724.DBW32634, 1 s

HMI tags "DB_SDC_ERROR_STAT_EMS071"
   "DB_SDC_ERRORS_STAT_ER_AKT[71].ER_TRIGER" : Word = PLC DB_SDC_ERRORS_STAT.ER_AKT[71].ER_TRIGER AT %DB3724.DBW32640, 1 s
   "DB_SDC_ERRORS_STAT_ER_AKT[71].ER_STAT[1].DRIVE_POS" : DInt = PLC DB_SDC_ERRORS_STAT.ER_AKT[71].ER_STAT[1].DRIVE_POS AT %DB3724.DBD32646, 1 s
   "DB_SDC_ERRORS_STAT_ER_AKT[71].ER_STAT[1].ERROR" : Int = PLC DB_SDC_ERRORS_STAT.ER_AKT[71].ER_STAT[1].ERROR AT %DB3724.DBW32652, 1 s
   "DB_SDC_ERRORS_STAT_ER_AKT[71].ER_STAT[2].DRIVE_POS" : DInt = PLC DB_SDC_ERRORS_STAT.ER_AKT[71].ER_STAT[2].DRIVE_POS AT %DB3724.DBD32662, 1 s
   "DB_SDC_ERRORS_STAT_ER_AKT[71].ER_STAT[2].ERROR" : Int = PLC DB_SDC_ERRORS_STAT.ER_AKT[71].ER_STAT[2].ERROR AT %DB3724.DBW32668, 1 s
   "DB_SDC_ERRORS_STAT_ER_AKT[71].ER_STAT[3].DRIVE_POS" : DInt = PLC DB_SDC_ERRORS_STAT.ER_AKT[71].ER_STAT[3].DRIVE_POS AT %DB3724.DBD32678, 1 s
   "DB_SDC_ERRORS_STAT_ER_AKT[71].ER_STAT[3].ERROR" : Int = PLC DB_SDC_ERRORS_STAT.ER_AKT[71].ER_STAT[3].ERROR AT %DB3724.DBW32684, 1 s
   "DB_SDC_ERRORS_STAT_ER_AKT[71].ER_STAT[4].DRIVE_POS" : DInt = PLC DB_SDC_ERRORS_STAT.ER_AKT[71].ER_STAT[4].DRIVE_POS AT %DB3724.DBD32694, 1 s
   "DB_SDC_ERRORS_STAT_ER_AKT[71].ER_STAT[4].ERROR" : Int = PLC DB_SDC_ERRORS_STAT.ER_AKT[71].ER_STAT[4].ERROR AT %DB3724.DBW32700, 1 s

HMI tags "DB_SDC_ERROR_STAT_EMS072"
   "DB_SDC_ERRORS_STAT_ER_AKT[72].ER_TRIGER" : Word = PLC DB_SDC_ERRORS_STAT.ER_AKT[72].ER_TRIGER AT %DB3724.DBW32706, 1 s
   "DB_SDC_ERRORS_STAT_ER_AKT[72].ER_STAT[1].DRIVE_POS" : DInt = PLC DB_SDC_ERRORS_STAT.ER_AKT[72].ER_STAT[1].DRIVE_POS AT %DB3724.DBD32712, 1 s
   "DB_SDC_ERRORS_STAT_ER_AKT[72].ER_STAT[1].ERROR" : Int = PLC DB_SDC_ERRORS_STAT.ER_AKT[72].ER_STAT[1].ERROR AT %DB3724.DBW32718, 1 s
   "DB_SDC_ERRORS_STAT_ER_AKT[72].ER_STAT[2].DRIVE_POS" : DInt = PLC DB_SDC_ERRORS_STAT.ER_AKT[72].ER_STAT[2].DRIVE_POS AT %DB3724.DBD32728, 1 s
   "DB_SDC_ERRORS_STAT_ER_AKT[72].ER_STAT[2].ERROR" : Int = PLC DB_SDC_ERRORS_STAT.ER_AKT[72].ER_STAT[2].ERROR AT %DB3724.DBW32734, 1 s
   "DB_SDC_ERRORS_STAT_ER_AKT[72].ER_STAT[3].DRIVE_POS" : DInt = PLC DB_SDC_ERRORS_STAT.ER_AKT[72].ER_STAT[3].DRIVE_POS AT %DB3724.DBD32744, 1 s
   "DB_SDC_ERRORS_STAT_ER_AKT[72].ER_STAT[3].ERROR" : Int = PLC DB_SDC_ERRORS_STAT.ER_AKT[72].ER_STAT[3].ERROR AT %DB3724.DBW32750, 1 s
   "DB_SDC_ERRORS_STAT_ER_AKT[72].ER_STAT[4].DRIVE_POS" : DInt = PLC DB_SDC_ERRORS_STAT.ER_AKT[72].ER_STAT[4].DRIVE_POS AT %DB3724.DBD32760, 1 s
   "DB_SDC_ERRORS_STAT_ER_AKT[72].ER_STAT[4].ERROR" : Int = PLC DB_SDC_ERRORS_STAT.ER_AKT[72].ER_STAT[4].ERROR AT %DB3724.DBW32766, 1 s

